REGION Network 6: IW210 - BWT Level (LT-422) - Tank #1
   RUNG wire#powerrail
      { S7_Templates := "[SrcType := Int, DestType := Real]" } Normalize(min := "20_TANKS_IP_DATA".RIO_03.FIRST_TANK.BWT_LEVEL_CNFG.RAW_MIN, value := "Tank 3P BWT Level", max := "20_TANKS_IP_DATA".RIO_03.FIRST_TANK.BWT_LEVEL_CNFG.RAW_MAX, out => "20_TANKS_IP_DATA".RIO_03.FIRST_TANK.BWT_LEVEL_CNFG.NORM)
      { S7_Templates := "[SrcType := Real, DestType := Real]" } Scale(min := "20_TANKS_IP_DATA".RIO_03.FIRST_TANK.BWT_LEVEL_CNFG.ENG_MIN, value := "IN_Level_WBT_3P", max := "20_TANKS_IP_DATA".RIO_03.FIRST_TANK.BWT_LEVEL_CNFG.ENG_MAX, out => "Tag_19")
      Move(in := "Data_From_WBT".Level_WBT_3P, out1 => "20_TANKS_IP_DATA".RIO_03.FIRST_TANK.BWT_LEVEL)
   END_RUNG
   // the same network as SCL:
   "20_TANKS_IP_DATA".RIO_03.FIRST_TANK.BWT_LEVEL_CNFG.NORM := NORM_X(MIN := "20_TANKS_IP_DATA".RIO_03.FIRST_TANK.BWT_LEVEL_CNFG.RAW_MIN, VALUE := "Tank 3P BWT Level", MAX := "20_TANKS_IP_DATA".RIO_03.FIRST_TANK.BWT_LEVEL_CNFG.RAW_MAX);
   "Tag_19" := SCALE_X(MIN := "20_TANKS_IP_DATA".RIO_03.FIRST_TANK.BWT_LEVEL_CNFG.ENG_MIN, VALUE := "IN_Level_WBT_3P", MAX := "20_TANKS_IP_DATA".RIO_03.FIRST_TANK.BWT_LEVEL_CNFG.ENG_MAX);
   "20_TANKS_IP_DATA".RIO_03.FIRST_TANK.BWT_LEVEL := "Data_From_WBT".Level_WBT_3P;
END_REGION

REGION Network 7: IW212 - BWT Level (LT-422) - Tank #2
   RUNG wire#powerrail
      { S7_Templates := "[SrcType := Int, DestType := Real]" } Normalize(min := "20_TANKS_IP_DATA".RIO_03.SECOND_TANK.BWT_LEVEL_CNFG.RAW_MIN, value := "Tank 3S BWT Level", max := "20_TANKS_IP_DATA".RIO_03.SECOND_TANK.BWT_LEVEL_CNFG.RAW_MAX, out => "20_TANKS_IP_DATA".RIO_03.SECOND_TANK.BWT_LEVEL_CNFG.NORM)
      { S7_Templates := "[SrcType := Real, DestType := Real]" } Scale(min := "20_TANKS_IP_DATA".RIO_03.SECOND_TANK.BWT_LEVEL_CNFG.ENG_MIN, value := "IN_Level_WBT_3S", max := "20_TANKS_IP_DATA".RIO_03.SECOND_TANK.BWT_LEVEL_CNFG.ENG_MAX, out => "Tag_21")
      Move(in := "Data_From_WBT".Level_WBT_3S, out1 => "20_TANKS_IP_DATA".RIO_03.SECOND_TANK.BWT_LEVEL)
   END_RUNG
   // the same network as SCL:
   "20_TANKS_IP_DATA".RIO_03.SECOND_TANK.BWT_LEVEL_CNFG.NORM := NORM_X(MIN := "20_TANKS_IP_DATA".RIO_03.SECOND_TANK.BWT_LEVEL_CNFG.RAW_MIN, VALUE := "Tank 3S BWT Level", MAX := "20_TANKS_IP_DATA".RIO_03.SECOND_TANK.BWT_LEVEL_CNFG.RAW_MAX);
   "Tag_21" := SCALE_X(MIN := "20_TANKS_IP_DATA".RIO_03.SECOND_TANK.BWT_LEVEL_CNFG.ENG_MIN, VALUE := "IN_Level_WBT_3S", MAX := "20_TANKS_IP_DATA".RIO_03.SECOND_TANK.BWT_LEVEL_CNFG.ENG_MAX);
   "20_TANKS_IP_DATA".RIO_03.SECOND_TANK.BWT_LEVEL := "Data_From_WBT".Level_WBT_3S;
END_REGION

REGION Network 8: IW214 - Spare Input - Tank #1
   RUNG wire#powerrail
      { S7_Templates := "[SrcType := Int, DestType := Real]" } Normalize(min := "20_TANKS_IP_DATA".RIO_03.FIRST_TANK.SPARE_AI_1_CNFG.RAW_MIN, value := "RIO3_SPR_AI_214", max := "20_TANKS_IP_DATA".RIO_03.FIRST_TANK.SPARE_AI_1_CNFG.RAW_MAX, out => "20_TANKS_IP_DATA".RIO_03.FIRST_TANK.SPARE_AI_1_CNFG.NORM)
      { S7_Templates := "[SrcType := Real, DestType := Real]" } Scale(min := "20_TANKS_IP_DATA".RIO_03.FIRST_TANK.SPARE_AI_1_CNFG.ENG_MIN, value := "20_TANKS_IP_DATA".RIO_03.FIRST_TANK.SPARE_AI_1_CNFG.NORM, max := "20_TANKS_IP_DATA".RIO_03.FIRST_TANK.SPARE_AI_1_CNFG.ENG_MAX, out => "20_TANKS_IP_DATA".RIO_03.FIRST_TANK.SPARE_AI_1)
   END_RUNG
   // the same network as SCL:
   "20_TANKS_IP_DATA".RIO_03.FIRST_TANK.SPARE_AI_1_CNFG.NORM := NORM_X(MIN := "20_TANKS_IP_DATA".RIO_03.FIRST_TANK.SPARE_AI_1_CNFG.RAW_MIN, VALUE := "RIO3_SPR_AI_214", MAX := "20_TANKS_IP_DATA".RIO_03.FIRST_TANK.SPARE_AI_1_CNFG.RAW_MAX);
   "20_TANKS_IP_DATA".RIO_03.FIRST_TANK.SPARE_AI_1 := SCALE_X(MIN := "20_TANKS_IP_DATA".RIO_03.FIRST_TANK.SPARE_AI_1_CNFG.ENG_MIN, VALUE := "20_TANKS_IP_DATA".RIO_03.FIRST_TANK.SPARE_AI_1_CNFG.NORM, MAX := "20_TANKS_IP_DATA".RIO_03.FIRST_TANK.SPARE_AI_1_CNFG.ENG_MAX);
END_REGION

REGION Network 9: IW216 - BWT Ph (426) - Tank #1
   RUNG wire#powerrail
      { S7_Templates := "[SrcType := Int, DestType := Real]" } Normalize(min := "20_TANKS_IP_DATA".RIO_03.FIRST_TANK.BWT_PH_CNFG.RAW_MIN, value := "Tank 3P BWT ph", max := "20_TANKS_IP_DATA".RIO_03.FIRST_TANK.BWT_PH_CNFG.RAW_MAX, out => "20_TANKS_IP_DATA".RIO_03.FIRST_TANK.BWT_PH_CNFG.NORM)
      { S7_Templates := "[SrcType := Real, DestType := Real]" } Scale(min := "20_TANKS_IP_DATA".RIO_03.FIRST_TANK.BWT_PH_CNFG.ENG_MIN, value := "20_TANKS_IP_DATA".RIO_03.FIRST_TANK.BWT_PH_CNFG.NORM, max := "20_TANKS_IP_DATA".RIO_03.FIRST_TANK.BWT_PH_CNFG.ENG_MAX, out => "20_TANKS_IP_DATA".RIO_03.FIRST_TANK.BWT_PH)
   END_RUNG
   // the same network as SCL:
   "20_TANKS_IP_DATA".RIO_03.FIRST_TANK.BWT_PH_CNFG.NORM := NORM_X(MIN := "20_TANKS_IP_DATA".RIO_03.FIRST_TANK.BWT_PH_CNFG.RAW_MIN, VALUE := "Tank 3P BWT ph", MAX := "20_TANKS_IP_DATA".RIO_03.FIRST_TANK.BWT_PH_CNFG.RAW_MAX);
   "20_TANKS_IP_DATA".RIO_03.FIRST_TANK.BWT_PH := SCALE_X(MIN := "20_TANKS_IP_DATA".RIO_03.FIRST_TANK.BWT_PH_CNFG.ENG_MIN, VALUE := "20_TANKS_IP_DATA".RIO_03.FIRST_TANK.BWT_PH_CNFG.NORM, MAX := "20_TANKS_IP_DATA".RIO_03.FIRST_TANK.BWT_PH_CNFG.ENG_MAX);
END_REGION

REGION Network 10: IW218 - BWT Temperature (426) - Tank #1
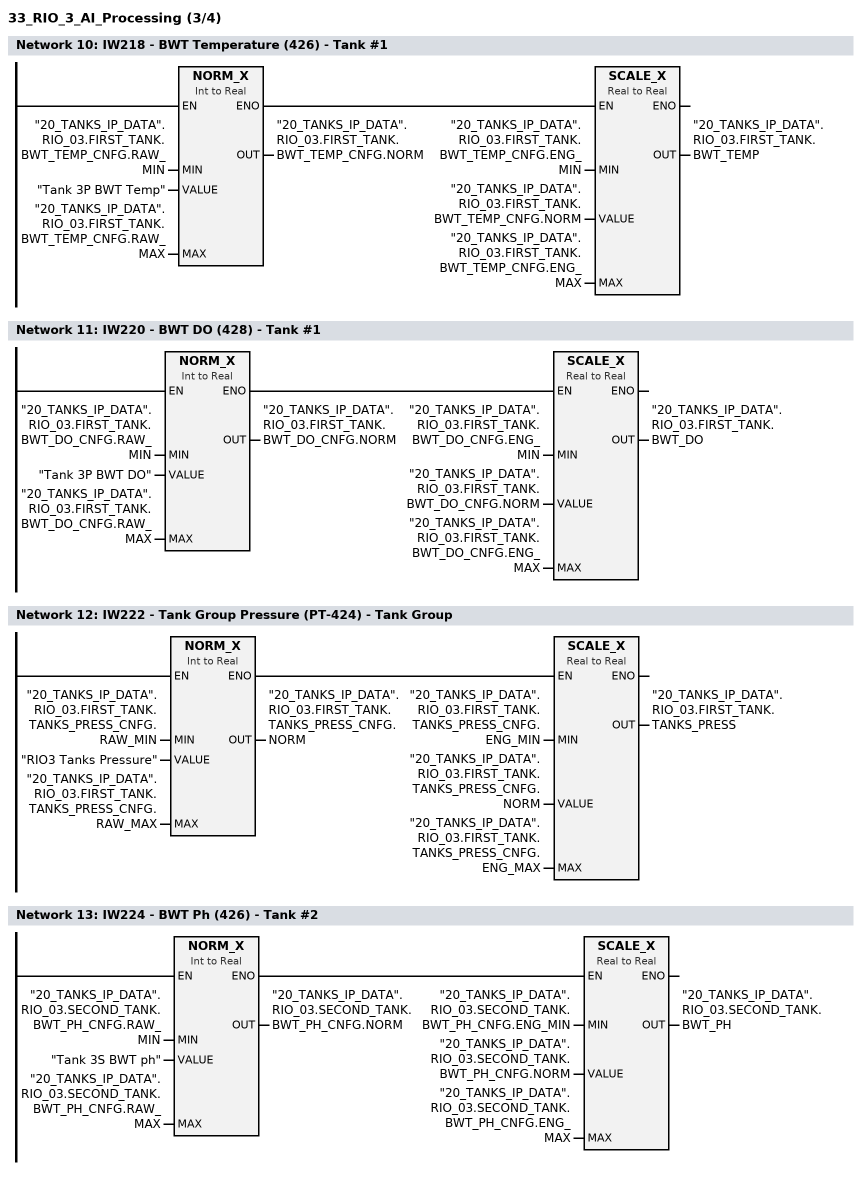
   RUNG wire#powerrail
      { S7_Templates := "[SrcType := Int, DestType := Real]" } Normalize(min := "20_TANKS_IP_DATA".RIO_03.FIRST_TANK.BWT_TEMP_CNFG.RAW_MIN, value := "Tank 3P BWT Temp", max := "20_TANKS_IP_DATA".RIO_03.FIRST_TANK.BWT_TEMP_CNFG.RAW_MAX, out => "20_TANKS_IP_DATA".RIO_03.FIRST_TANK.BWT_TEMP_CNFG.NORM)
      { S7_Templates := "[SrcType := Real, DestType := Real]" } Scale(min := "20_TANKS_IP_DATA".RIO_03.FIRST_TANK.BWT_TEMP_CNFG.ENG_MIN, value := "20_TANKS_IP_DATA".RIO_03.FIRST_TANK.BWT_TEMP_CNFG.NORM, max := "20_TANKS_IP_DATA".RIO_03.FIRST_TANK.BWT_TEMP_CNFG.ENG_MAX, out => "20_TANKS_IP_DATA".RIO_03.FIRST_TANK.BWT_TEMP)
   END_RUNG
   // the same network as SCL:
   "20_TANKS_IP_DATA".RIO_03.FIRST_TANK.BWT_TEMP_CNFG.NORM := NORM_X(MIN := "20_TANKS_IP_DATA".RIO_03.FIRST_TANK.BWT_TEMP_CNFG.RAW_MIN, VALUE := "Tank 3P BWT Temp", MAX := "20_TANKS_IP_DATA".RIO_03.FIRST_TANK.BWT_TEMP_CNFG.RAW_MAX);
   "20_TANKS_IP_DATA".RIO_03.FIRST_TANK.BWT_TEMP := SCALE_X(MIN := "20_TANKS_IP_DATA".RIO_03.FIRST_TANK.BWT_TEMP_CNFG.ENG_MIN, VALUE := "20_TANKS_IP_DATA".RIO_03.FIRST_TANK.BWT_TEMP_CNFG.NORM, MAX := "20_TANKS_IP_DATA".RIO_03.FIRST_TANK.BWT_TEMP_CNFG.ENG_MAX);
END_REGION

REGION Network 11: IW220 - BWT DO (428) - Tank #1
   RUNG wire#powerrail
      { S7_Templates := "[SrcType := Int, DestType := Real]" } Normalize(min := "20_TANKS_IP_DATA".RIO_03.FIRST_TANK.BWT_DO_CNFG.RAW_MIN, value := "Tank 3P BWT DO", max := "20_TANKS_IP_DATA".RIO_03.FIRST_TANK.BWT_DO_CNFG.RAW_MAX, out => "20_TANKS_IP_DATA".RIO_03.FIRST_TANK.BWT_DO_CNFG.NORM)
      { S7_Templates := "[SrcType := Real, DestType := Real]" } Scale(min := "20_TANKS_IP_DATA".RIO_03.FIRST_TANK.BWT_DO_CNFG.ENG_MIN, value := "20_TANKS_IP_DATA".RIO_03.FIRST_TANK.BWT_DO_CNFG.NORM, max := "20_TANKS_IP_DATA".RIO_03.FIRST_TANK.BWT_DO_CNFG.ENG_MAX, out => "20_TANKS_IP_DATA".RIO_03.FIRST_TANK.BWT_DO)
   END_RUNG
   // the same network as SCL:
   "20_TANKS_IP_DATA".RIO_03.FIRST_TANK.BWT_DO_CNFG.NORM := NORM_X(MIN := "20_TANKS_IP_DATA".RIO_03.FIRST_TANK.BWT_DO_CNFG.RAW_MIN, VALUE := "Tank 3P BWT DO", MAX := "20_TANKS_IP_DATA".RIO_03.FIRST_TANK.BWT_DO_CNFG.RAW_MAX);
   "20_TANKS_IP_DATA".RIO_03.FIRST_TANK.BWT_DO := SCALE_X(MIN := "20_TANKS_IP_DATA".RIO_03.FIRST_TANK.BWT_DO_CNFG.ENG_MIN, VALUE := "20_TANKS_IP_DATA".RIO_03.FIRST_TANK.BWT_DO_CNFG.NORM, MAX := "20_TANKS_IP_DATA".RIO_03.FIRST_TANK.BWT_DO_CNFG.ENG_MAX);
END_REGION

REGION Network 12: IW222 - Tank Group Pressure (PT-424) - Tank Group
   RUNG wire#powerrail
      { S7_Templates := "[SrcType := Int, DestType := Real]" } Normalize(min := "20_TANKS_IP_DATA".RIO_03.FIRST_TANK.TANKS_PRESS_CNFG.RAW_MIN, value := "RIO3 Tanks Pressure", max := "20_TANKS_IP_DATA".RIO_03.FIRST_TANK.TANKS_PRESS_CNFG.RAW_MAX, out => "20_TANKS_IP_DATA".RIO_03.FIRST_TANK.TANKS_PRESS_CNFG.NORM)
      { S7_Templates := "[SrcType := Real, DestType := Real]" } Scale(min := "20_TANKS_IP_DATA".RIO_03.FIRST_TANK.TANKS_PRESS_CNFG.ENG_MIN, value := "20_TANKS_IP_DATA".RIO_03.FIRST_TANK.TANKS_PRESS_CNFG.NORM, max := "20_TANKS_IP_DATA".RIO_03.FIRST_TANK.TANKS_PRESS_CNFG.ENG_MAX, out => "20_TANKS_IP_DATA".RIO_03.FIRST_TANK.TANKS_PRESS)
   END_RUNG
   // the same network as SCL:
   "20_TANKS_IP_DATA".RIO_03.FIRST_TANK.TANKS_PRESS_CNFG.NORM := NORM_X(MIN := "20_TANKS_IP_DATA".RIO_03.FIRST_TANK.TANKS_PRESS_CNFG.RAW_MIN, VALUE := "RIO3 Tanks Pressure", MAX := "20_TANKS_IP_DATA".RIO_03.FIRST_TANK.TANKS_PRESS_CNFG.RAW_MAX);
   "20_TANKS_IP_DATA".RIO_03.FIRST_TANK.TANKS_PRESS := SCALE_X(MIN := "20_TANKS_IP_DATA".RIO_03.FIRST_TANK.TANKS_PRESS_CNFG.ENG_MIN, VALUE := "20_TANKS_IP_DATA".RIO_03.FIRST_TANK.TANKS_PRESS_CNFG.NORM, MAX := "20_TANKS_IP_DATA".RIO_03.FIRST_TANK.TANKS_PRESS_CNFG.ENG_MAX);
END_REGION

REGION Network 13: IW224 - BWT Ph (426) - Tank #2
   RUNG wire#powerrail
      { S7_Templates := "[SrcType := Int, DestType := Real]" } Normalize(min := "20_TANKS_IP_DATA".RIO_03.SECOND_TANK.BWT_PH_CNFG.RAW_MIN, value := "Tank 3S BWT ph", max := "20_TANKS_IP_DATA".RIO_03.SECOND_TANK.BWT_PH_CNFG.RAW_MAX, out => "20_TANKS_IP_DATA".RIO_03.SECOND_TANK.BWT_PH_CNFG.NORM)
      { S7_Templates := "[SrcType := Real, DestType := Real]" } Scale(min := "20_TANKS_IP_DATA".RIO_03.SECOND_TANK.BWT_PH_CNFG.ENG_MIN, value := "20_TANKS_IP_DATA".RIO_03.SECOND_TANK.BWT_PH_CNFG.NORM, max := "20_TANKS_IP_DATA".RIO_03.SECOND_TANK.BWT_PH_CNFG.ENG_MAX, out => "20_TANKS_IP_DATA".RIO_03.SECOND_TANK.BWT_PH)
   END_RUNG
   // the same network as SCL:
   "20_TANKS_IP_DATA".RIO_03.SECOND_TANK.BWT_PH_CNFG.NORM := NORM_X(MIN := "20_TANKS_IP_DATA".RIO_03.SECOND_TANK.BWT_PH_CNFG.RAW_MIN, VALUE := "Tank 3S BWT ph", MAX := "20_TANKS_IP_DATA".RIO_03.SECOND_TANK.BWT_PH_CNFG.RAW_MAX);
   "20_TANKS_IP_DATA".RIO_03.SECOND_TANK.BWT_PH := SCALE_X(MIN := "20_TANKS_IP_DATA".RIO_03.SECOND_TANK.BWT_PH_CNFG.ENG_MIN, VALUE := "20_TANKS_IP_DATA".RIO_03.SECOND_TANK.BWT_PH_CNFG.NORM, MAX := "20_TANKS_IP_DATA".RIO_03.SECOND_TANK.BWT_PH_CNFG.ENG_MAX);
END_REGION

REGION Network 14: IW226 - BWT Temperature (426) - Tank #2
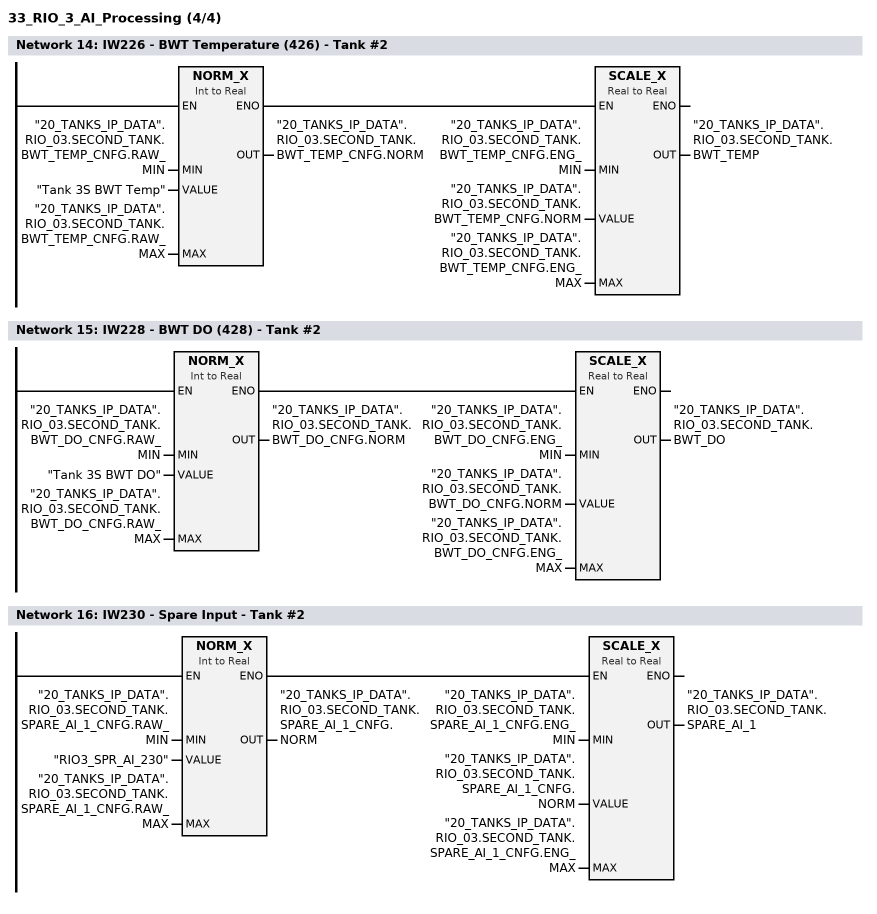
   RUNG wire#powerrail
      { S7_Templates := "[SrcType := Int, DestType := Real]" } Normalize(min := "20_TANKS_IP_DATA".RIO_03.SECOND_TANK.BWT_TEMP_CNFG.RAW_MIN, value := "Tank 3S BWT Temp", max := "20_TANKS_IP_DATA".RIO_03.SECOND_TANK.BWT_TEMP_CNFG.RAW_MAX, out => "20_TANKS_IP_DATA".RIO_03.SECOND_TANK.BWT_TEMP_CNFG.NORM)
      { S7_Templates := "[SrcType := Real, DestType := Real]" } Scale(min := "20_TANKS_IP_DATA".RIO_03.SECOND_TANK.BWT_TEMP_CNFG.ENG_MIN, value := "20_TANKS_IP_DATA".RIO_03.SECOND_TANK.BWT_TEMP_CNFG.NORM, max := "20_TANKS_IP_DATA".RIO_03.SECOND_TANK.BWT_TEMP_CNFG.ENG_MAX, out => "20_TANKS_IP_DATA".RIO_03.SECOND_TANK.BWT_TEMP)
   END_RUNG
   // the same network as SCL:
   "20_TANKS_IP_DATA".RIO_03.SECOND_TANK.BWT_TEMP_CNFG.NORM := NORM_X(MIN := "20_TANKS_IP_DATA".RIO_03.SECOND_TANK.BWT_TEMP_CNFG.RAW_MIN, VALUE := "Tank 3S BWT Temp", MAX := "20_TANKS_IP_DATA".RIO_03.SECOND_TANK.BWT_TEMP_CNFG.RAW_MAX);
   "20_TANKS_IP_DATA".RIO_03.SECOND_TANK.BWT_TEMP := SCALE_X(MIN := "20_TANKS_IP_DATA".RIO_03.SECOND_TANK.BWT_TEMP_CNFG.ENG_MIN, VALUE := "20_TANKS_IP_DATA".RIO_03.SECOND_TANK.BWT_TEMP_CNFG.NORM, MAX := "20_TANKS_IP_DATA".RIO_03.SECOND_TANK.BWT_TEMP_CNFG.ENG_MAX);
END_REGION

REGION Network 15: IW228 - BWT DO (428) - Tank #2
   RUNG wire#powerrail
      { S7_Templates := "[SrcType := Int, DestType := Real]" } Normalize(min := "20_TANKS_IP_DATA".RIO_03.SECOND_TANK.BWT_DO_CNFG.RAW_MIN, value := "Tank 3S BWT DO", max := "20_TANKS_IP_DATA".RIO_03.SECOND_TANK.BWT_DO_CNFG.RAW_MAX, out => "20_TANKS_IP_DATA".RIO_03.SECOND_TANK.BWT_DO_CNFG.NORM)
      { S7_Templates := "[SrcType := Real, DestType := Real]" } Scale(min := "20_TANKS_IP_DATA".RIO_03.SECOND_TANK.BWT_DO_CNFG.ENG_MIN, value := "20_TANKS_IP_DATA".RIO_03.SECOND_TANK.BWT_DO_CNFG.NORM, max := "20_TANKS_IP_DATA".RIO_03.SECOND_TANK.BWT_DO_CNFG.ENG_MAX, out => "20_TANKS_IP_DATA".RIO_03.SECOND_TANK.BWT_DO)
   END_RUNG
   // the same network as SCL:
   "20_TANKS_IP_DATA".RIO_03.SECOND_TANK.BWT_DO_CNFG.NORM := NORM_X(MIN := "20_TANKS_IP_DATA".RIO_03.SECOND_TANK.BWT_DO_CNFG.RAW_MIN, VALUE := "Tank 3S BWT DO", MAX := "20_TANKS_IP_DATA".RIO_03.SECOND_TANK.BWT_DO_CNFG.RAW_MAX);
   "20_TANKS_IP_DATA".RIO_03.SECOND_TANK.BWT_DO := SCALE_X(MIN := "20_TANKS_IP_DATA".RIO_03.SECOND_TANK.BWT_DO_CNFG.ENG_MIN, VALUE := "20_TANKS_IP_DATA".RIO_03.SECOND_TANK.BWT_DO_CNFG.NORM, MAX := "20_TANKS_IP_DATA".RIO_03.SECOND_TANK.BWT_DO_CNFG.ENG_MAX);
END_REGION

REGION Network 16: IW230 - Spare Input - Tank #2
   RUNG wire#powerrail
      { S7_Templates := "[SrcType := Int, DestType := Real]" } Normalize(min := "20_TANKS_IP_DATA".RIO_03.SECOND_TANK.SPARE_AI_1_CNFG.RAW_MIN, value := "RIO3_SPR_AI_230", max := "20_TANKS_IP_DATA".RIO_03.SECOND_TANK.SPARE_AI_1_CNFG.RAW_MAX, out => "20_TANKS_IP_DATA".RIO_03.SECOND_TANK.SPARE_AI_1_CNFG.NORM)
      { S7_Templates := "[SrcType := Real, DestType := Real]" } Scale(min := "20_TANKS_IP_DATA".RIO_03.SECOND_TANK.SPARE_AI_1_CNFG.ENG_MIN, value := "20_TANKS_IP_DATA".RIO_03.SECOND_TANK.SPARE_AI_1_CNFG.NORM, max := "20_TANKS_IP_DATA".RIO_03.SECOND_TANK.SPARE_AI_1_CNFG.ENG_MAX, out => "20_TANKS_IP_DATA".RIO_03.SECOND_TANK.SPARE_AI_1)
   END_RUNG
   // the same network as SCL:
   "20_TANKS_IP_DATA".RIO_03.SECOND_TANK.SPARE_AI_1_CNFG.NORM := NORM_X(MIN := "20_TANKS_IP_DATA".RIO_03.SECOND_TANK.SPARE_AI_1_CNFG.RAW_MIN, VALUE := "RIO3_SPR_AI_230", MAX := "20_TANKS_IP_DATA".RIO_03.SECOND_TANK.SPARE_AI_1_CNFG.RAW_MAX);
   "20_TANKS_IP_DATA".RIO_03.SECOND_TANK.SPARE_AI_1 := SCALE_X(MIN := "20_TANKS_IP_DATA".RIO_03.SECOND_TANK.SPARE_AI_1_CNFG.ENG_MIN, VALUE := "20_TANKS_IP_DATA".RIO_03.SECOND_TANK.SPARE_AI_1_CNFG.NORM, MAX := "20_TANKS_IP_DATA".RIO_03.SECOND_TANK.SPARE_AI_1_CNFG.ENG_MAX);
END_REGION
END_FUNCTION

FUNCTION "34_RIO_4_AI_Processing" : Void   // FC34, LAD
TITLE = Analogue Input Processing (Tank 1 = 4P, Tank 2 = 4S)
{ S7_Optimized_Access := 'TRUE' }
AUTHOR : JRS
VERSION : 0.1
// To process raw inputs prior to code use
BEGIN

REGION Network 1: IW260 - USD Flow (FIT-418) - Tank #1
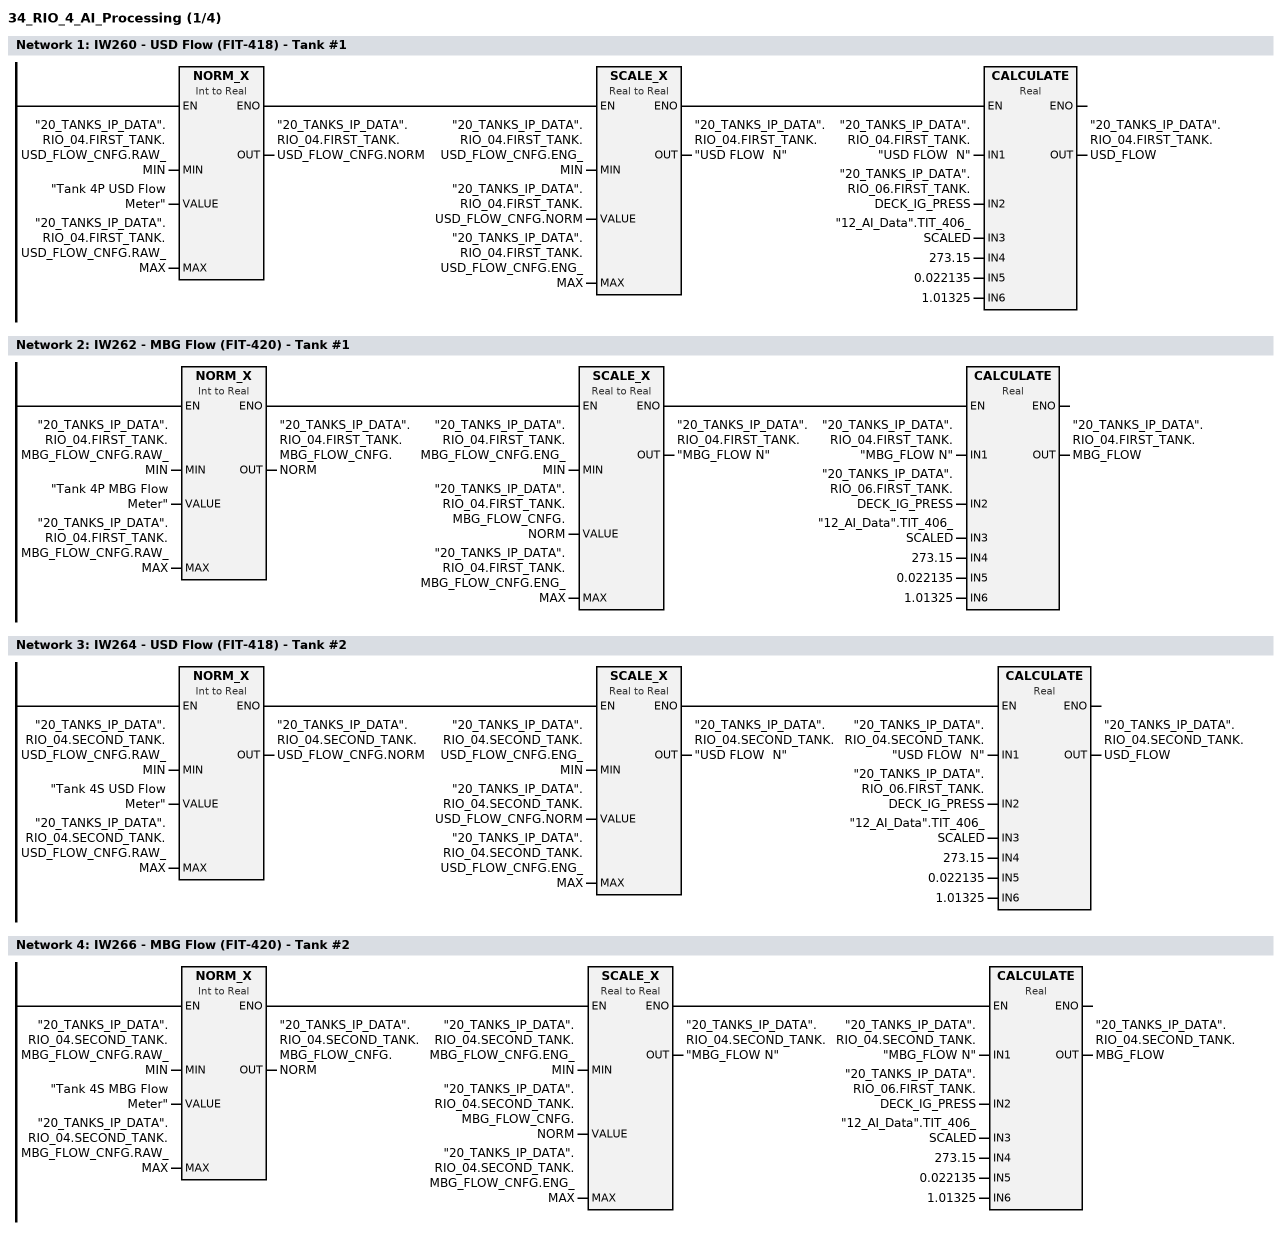
   RUNG wire#powerrail
      { S7_Templates := "[SrcType := Int, DestType := Real]" } Normalize(min := "20_TANKS_IP_DATA".RIO_04.FIRST_TANK.USD_FLOW_CNFG.RAW_MIN, value := "Tank 4P USD Flow Meter", max := "20_TANKS_IP_DATA".RIO_04.FIRST_TANK.USD_FLOW_CNFG.RAW_MAX, out => "20_TANKS_IP_DATA".RIO_04.FIRST_TANK.USD_FLOW_CNFG.NORM)
      { S7_Templates := "[SrcType := Real, DestType := Real]" } Scale(min := "20_TANKS_IP_DATA".RIO_04.FIRST_TANK.USD_FLOW_CNFG.ENG_MIN, value := "20_TANKS_IP_DATA".RIO_04.FIRST_TANK.USD_FLOW_CNFG.NORM, max := "20_TANKS_IP_DATA".RIO_04.FIRST_TANK.USD_FLOW_CNFG.ENG_MAX, out => "20_TANKS_IP_DATA".RIO_04.FIRST_TANK."USD FLOW  N")
      { S7_Templates := "SrcType := Real"; S7_Expression := "IN1*(IN2+IN6)/IN6*IN4/(IN3+IN4)" } Calculate(in1 := "20_TANKS_IP_DATA".RIO_04.FIRST_TANK."USD FLOW  N", in2 := "20_TANKS_IP_DATA".RIO_06.FIRST_TANK.DECK_IG_PRESS, in3 := "12_AI_Data".TIT_406_SCALED, in4 := 273.15, in5 := 0.022135, in6 := 1.01325, out => "20_TANKS_IP_DATA".RIO_04.FIRST_TANK.USD_FLOW)
   END_RUNG
   // the same network as SCL:
   "20_TANKS_IP_DATA".RIO_04.FIRST_TANK.USD_FLOW_CNFG.NORM := NORM_X(MIN := "20_TANKS_IP_DATA".RIO_04.FIRST_TANK.USD_FLOW_CNFG.RAW_MIN, VALUE := "Tank 4P USD Flow Meter", MAX := "20_TANKS_IP_DATA".RIO_04.FIRST_TANK.USD_FLOW_CNFG.RAW_MAX);
   "20_TANKS_IP_DATA".RIO_04.FIRST_TANK."USD FLOW  N" := SCALE_X(MIN := "20_TANKS_IP_DATA".RIO_04.FIRST_TANK.USD_FLOW_CNFG.ENG_MIN, VALUE := "20_TANKS_IP_DATA".RIO_04.FIRST_TANK.USD_FLOW_CNFG.NORM, MAX := "20_TANKS_IP_DATA".RIO_04.FIRST_TANK.USD_FLOW_CNFG.ENG_MAX);
   "20_TANKS_IP_DATA".RIO_04.FIRST_TANK.USD_FLOW := "20_TANKS_IP_DATA".RIO_04.FIRST_TANK."USD FLOW  N"*("20_TANKS_IP_DATA".RIO_06.FIRST_TANK.DECK_IG_PRESS+1.01325)/1.01325*273.15/("12_AI_Data".TIT_406_SCALED+273.15);
END_REGION

REGION Network 2: IW262 - MBG Flow (FIT-420) - Tank #1
   RUNG wire#powerrail
      { S7_Templates := "[SrcType := Int, DestType := Real]" } Normalize(min := "20_TANKS_IP_DATA".RIO_04.FIRST_TANK.MBG_FLOW_CNFG.RAW_MIN, value := "Tank 4P MBG Flow Meter", max := "20_TANKS_IP_DATA".RIO_04.FIRST_TANK.MBG_FLOW_CNFG.RAW_MAX, out => "20_TANKS_IP_DATA".RIO_04.FIRST_TANK.MBG_FLOW_CNFG.NORM)
      { S7_Templates := "[SrcType := Real, DestType := Real]" } Scale(min := "20_TANKS_IP_DATA".RIO_04.FIRST_TANK.MBG_FLOW_CNFG.ENG_MIN, value := "20_TANKS_IP_DATA".RIO_04.FIRST_TANK.MBG_FLOW_CNFG.NORM, max := "20_TANKS_IP_DATA".RIO_04.FIRST_TANK.MBG_FLOW_CNFG.ENG_MAX, out => "20_TANKS_IP_DATA".RIO_04.FIRST_TANK."MBG_FLOW N")
      { S7_Templates := "SrcType := Real"; S7_Expression := "IN1*(IN2+IN6)/IN6*IN4/(IN3+IN4)" } Calculate(in1 := "20_TANKS_IP_DATA".RIO_04.FIRST_TANK."MBG_FLOW N", in2 := "20_TANKS_IP_DATA".RIO_06.FIRST_TANK.DECK_IG_PRESS, in3 := "12_AI_Data".TIT_406_SCALED, in4 := 273.15, in5 := 0.022135, in6 := 1.01325, out => "20_TANKS_IP_DATA".RIO_04.FIRST_TANK.MBG_FLOW)
   END_RUNG
   // the same network as SCL:
   "20_TANKS_IP_DATA".RIO_04.FIRST_TANK.MBG_FLOW_CNFG.NORM := NORM_X(MIN := "20_TANKS_IP_DATA".RIO_04.FIRST_TANK.MBG_FLOW_CNFG.RAW_MIN, VALUE := "Tank 4P MBG Flow Meter", MAX := "20_TANKS_IP_DATA".RIO_04.FIRST_TANK.MBG_FLOW_CNFG.RAW_MAX);
   "20_TANKS_IP_DATA".RIO_04.FIRST_TANK."MBG_FLOW N" := SCALE_X(MIN := "20_TANKS_IP_DATA".RIO_04.FIRST_TANK.MBG_FLOW_CNFG.ENG_MIN, VALUE := "20_TANKS_IP_DATA".RIO_04.FIRST_TANK.MBG_FLOW_CNFG.NORM, MAX := "20_TANKS_IP_DATA".RIO_04.FIRST_TANK.MBG_FLOW_CNFG.ENG_MAX);
   "20_TANKS_IP_DATA".RIO_04.FIRST_TANK.MBG_FLOW := "20_TANKS_IP_DATA".RIO_04.FIRST_TANK."MBG_FLOW N"*("20_TANKS_IP_DATA".RIO_06.FIRST_TANK.DECK_IG_PRESS+1.01325)/1.01325*273.15/("12_AI_Data".TIT_406_SCALED+273.15);
END_REGION

REGION Network 3: IW264 - USD Flow (FIT-418) - Tank #2
   RUNG wire#powerrail
      { S7_Templates := "[SrcType := Int, DestType := Real]" } Normalize(min := "20_TANKS_IP_DATA".RIO_04.SECOND_TANK.USD_FLOW_CNFG.RAW_MIN, value := "Tank 4S USD Flow Meter", max := "20_TANKS_IP_DATA".RIO_04.SECOND_TANK.USD_FLOW_CNFG.RAW_MAX, out => "20_TANKS_IP_DATA".RIO_04.SECOND_TANK.USD_FLOW_CNFG.NORM)
      { S7_Templates := "[SrcType := Real, DestType := Real]" } Scale(min := "20_TANKS_IP_DATA".RIO_04.SECOND_TANK.USD_FLOW_CNFG.ENG_MIN, value := "20_TANKS_IP_DATA".RIO_04.SECOND_TANK.USD_FLOW_CNFG.NORM, max := "20_TANKS_IP_DATA".RIO_04.SECOND_TANK.USD_FLOW_CNFG.ENG_MAX, out => "20_TANKS_IP_DATA".RIO_04.SECOND_TANK."USD FLOW  N")
      { S7_Templates := "SrcType := Real"; S7_Expression := "IN1*(IN2+IN6)/IN6*IN4/(IN3+IN4)" } Calculate(in1 := "20_TANKS_IP_DATA".RIO_04.SECOND_TANK."USD FLOW  N", in2 := "20_TANKS_IP_DATA".RIO_06.FIRST_TANK.DECK_IG_PRESS, in3 := "12_AI_Data".TIT_406_SCALED, in4 := 273.15, in5 := 0.022135, in6 := 1.01325, out => "20_TANKS_IP_DATA".RIO_04.SECOND_TANK.USD_FLOW)
   END_RUNG
   // the same network as SCL:
   "20_TANKS_IP_DATA".RIO_04.SECOND_TANK.USD_FLOW_CNFG.NORM := NORM_X(MIN := "20_TANKS_IP_DATA".RIO_04.SECOND_TANK.USD_FLOW_CNFG.RAW_MIN, VALUE := "Tank 4S USD Flow Meter", MAX := "20_TANKS_IP_DATA".RIO_04.SECOND_TANK.USD_FLOW_CNFG.RAW_MAX);
   "20_TANKS_IP_DATA".RIO_04.SECOND_TANK."USD FLOW  N" := SCALE_X(MIN := "20_TANKS_IP_DATA".RIO_04.SECOND_TANK.USD_FLOW_CNFG.ENG_MIN, VALUE := "20_TANKS_IP_DATA".RIO_04.SECOND_TANK.USD_FLOW_CNFG.NORM, MAX := "20_TANKS_IP_DATA".RIO_04.SECOND_TANK.USD_FLOW_CNFG.ENG_MAX);
   "20_TANKS_IP_DATA".RIO_04.SECOND_TANK.USD_FLOW := "20_TANKS_IP_DATA".RIO_04.SECOND_TANK."USD FLOW  N"*("20_TANKS_IP_DATA".RIO_06.FIRST_TANK.DECK_IG_PRESS+1.01325)/1.01325*273.15/("12_AI_Data".TIT_406_SCALED+273.15);
END_REGION

REGION Network 4: IW266 - MBG Flow (FIT-420) - Tank #2
   RUNG wire#powerrail
      { S7_Templates := "[SrcType := Int, DestType := Real]" } Normalize(min := "20_TANKS_IP_DATA".RIO_04.SECOND_TANK.MBG_FLOW_CNFG.RAW_MIN, value := "Tank 4S MBG Flow Meter", max := "20_TANKS_IP_DATA".RIO_04.SECOND_TANK.MBG_FLOW_CNFG.RAW_MAX, out => "20_TANKS_IP_DATA".RIO_04.SECOND_TANK.MBG_FLOW_CNFG.NORM)
      { S7_Templates := "[SrcType := Real, DestType := Real]" } Scale(min := "20_TANKS_IP_DATA".RIO_04.SECOND_TANK.MBG_FLOW_CNFG.ENG_MIN, value := "20_TANKS_IP_DATA".RIO_04.SECOND_TANK.MBG_FLOW_CNFG.NORM, max := "20_TANKS_IP_DATA".RIO_04.SECOND_TANK.MBG_FLOW_CNFG.ENG_MAX, out => "20_TANKS_IP_DATA".RIO_04.SECOND_TANK."MBG_FLOW N")
      { S7_Templates := "SrcType := Real"; S7_Expression := "IN1*(IN2+IN6)/IN6*IN4/(IN3+IN4)" } Calculate(in1 := "20_TANKS_IP_DATA".RIO_04.SECOND_TANK."MBG_FLOW N", in2 := "20_TANKS_IP_DATA".RIO_06.FIRST_TANK.DECK_IG_PRESS, in3 := "12_AI_Data".TIT_406_SCALED, in4 := 273.15, in5 := 0.022135, in6 := 1.01325, out => "20_TANKS_IP_DATA".RIO_04.SECOND_TANK.MBG_FLOW)
   END_RUNG
   // the same network as SCL:
   "20_TANKS_IP_DATA".RIO_04.SECOND_TANK.MBG_FLOW_CNFG.NORM := NORM_X(MIN := "20_TANKS_IP_DATA".RIO_04.SECOND_TANK.MBG_FLOW_CNFG.RAW_MIN, VALUE := "Tank 4S MBG Flow Meter", MAX := "20_TANKS_IP_DATA".RIO_04.SECOND_TANK.MBG_FLOW_CNFG.RAW_MAX);
   "20_TANKS_IP_DATA".RIO_04.SECOND_TANK."MBG_FLOW N" := SCALE_X(MIN := "20_TANKS_IP_DATA".RIO_04.SECOND_TANK.MBG_FLOW_CNFG.ENG_MIN, VALUE := "20_TANKS_IP_DATA".RIO_04.SECOND_TANK.MBG_FLOW_CNFG.NORM, MAX := "20_TANKS_IP_DATA".RIO_04.SECOND_TANK.MBG_FLOW_CNFG.ENG_MAX);
   "20_TANKS_IP_DATA".RIO_04.SECOND_TANK.MBG_FLOW := "20_TANKS_IP_DATA".RIO_04.SECOND_TANK."MBG_FLOW N"*("20_TANKS_IP_DATA".RIO_06.FIRST_TANK.DECK_IG_PRESS+1.01325)/1.01325*273.15/("12_AI_Data".TIT_406_SCALED+273.15);
END_REGION

REGION Network 5: IW268 - Deck Main IG Pressure (PT-415) - Tank Group
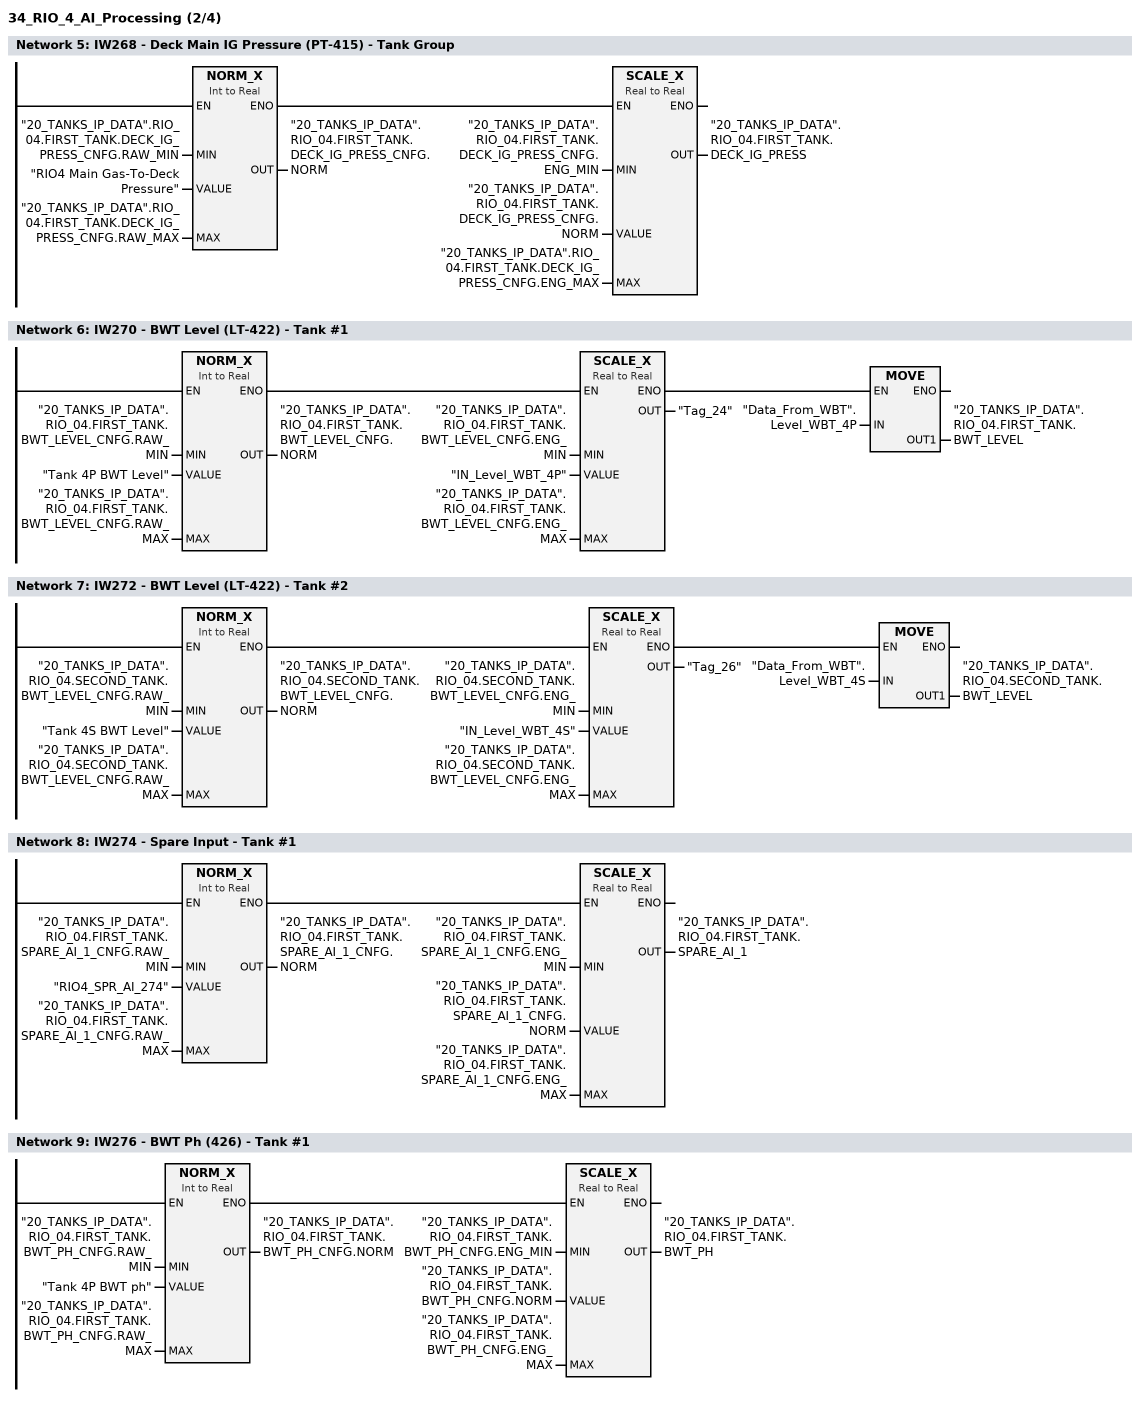
   RUNG wire#powerrail
      { S7_Templates := "[SrcType := Int, DestType := Real]" } Normalize(min := "20_TANKS_IP_DATA".RIO_04.FIRST_TANK.DECK_IG_PRESS_CNFG.RAW_MIN, value := "RIO4 Main Gas-To-Deck Pressure", max := "20_TANKS_IP_DATA".RIO_04.FIRST_TANK.DECK_IG_PRESS_CNFG.RAW_MAX, out => "20_TANKS_IP_DATA".RIO_04.FIRST_TANK.DECK_IG_PRESS_CNFG.NORM)
      { S7_Templates := "[SrcType := Real, DestType := Real]" } Scale(min := "20_TANKS_IP_DATA".RIO_04.FIRST_TANK.DECK_IG_PRESS_CNFG.ENG_MIN, value := "20_TANKS_IP_DATA".RIO_04.FIRST_TANK.DECK_IG_PRESS_CNFG.NORM, max := "20_TANKS_IP_DATA".RIO_04.FIRST_TANK.DECK_IG_PRESS_CNFG.ENG_MAX, out => "20_TANKS_IP_DATA".RIO_04.FIRST_TANK.DECK_IG_PRESS)
   END_RUNG
   // the same network as SCL:
   "20_TANKS_IP_DATA".RIO_04.FIRST_TANK.DECK_IG_PRESS_CNFG.NORM := NORM_X(MIN := "20_TANKS_IP_DATA".RIO_04.FIRST_TANK.DECK_IG_PRESS_CNFG.RAW_MIN, VALUE := "RIO4 Main Gas-To-Deck Pressure", MAX := "20_TANKS_IP_DATA".RIO_04.FIRST_TANK.DECK_IG_PRESS_CNFG.RAW_MAX);
   "20_TANKS_IP_DATA".RIO_04.FIRST_TANK.DECK_IG_PRESS := SCALE_X(MIN := "20_TANKS_IP_DATA".RIO_04.FIRST_TANK.DECK_IG_PRESS_CNFG.ENG_MIN, VALUE := "20_TANKS_IP_DATA".RIO_04.FIRST_TANK.DECK_IG_PRESS_CNFG.NORM, MAX := "20_TANKS_IP_DATA".RIO_04.FIRST_TANK.DECK_IG_PRESS_CNFG.ENG_MAX);
END_REGION

REGION Network 6: IW270 - BWT Level (LT-422) - Tank #1
   RUNG wire#powerrail
      { S7_Templates := "[SrcType := Int, DestType := Real]" } Normalize(min := "20_TANKS_IP_DATA".RIO_04.FIRST_TANK.BWT_LEVEL_CNFG.RAW_MIN, value := "Tank 4P BWT Level", max := "20_TANKS_IP_DATA".RIO_04.FIRST_TANK.BWT_LEVEL_CNFG.RAW_MAX, out => "20_TANKS_IP_DATA".RIO_04.FIRST_TANK.BWT_LEVEL_CNFG.NORM)
      { S7_Templates := "[SrcType := Real, DestType := Real]" } Scale(min := "20_TANKS_IP_DATA".RIO_04.FIRST_TANK.BWT_LEVEL_CNFG.ENG_MIN, value := "IN_Level_WBT_4P", max := "20_TANKS_IP_DATA".RIO_04.FIRST_TANK.BWT_LEVEL_CNFG.ENG_MAX, out => "Tag_24")
      Move(in := "Data_From_WBT".Level_WBT_4P, out1 => "20_TANKS_IP_DATA".RIO_04.FIRST_TANK.BWT_LEVEL)
   END_RUNG
   // the same network as SCL:
   "20_TANKS_IP_DATA".RIO_04.FIRST_TANK.BWT_LEVEL_CNFG.NORM := NORM_X(MIN := "20_TANKS_IP_DATA".RIO_04.FIRST_TANK.BWT_LEVEL_CNFG.RAW_MIN, VALUE := "Tank 4P BWT Level", MAX := "20_TANKS_IP_DATA".RIO_04.FIRST_TANK.BWT_LEVEL_CNFG.RAW_MAX);
   "Tag_24" := SCALE_X(MIN := "20_TANKS_IP_DATA".RIO_04.FIRST_TANK.BWT_LEVEL_CNFG.ENG_MIN, VALUE := "IN_Level_WBT_4P", MAX := "20_TANKS_IP_DATA".RIO_04.FIRST_TANK.BWT_LEVEL_CNFG.ENG_MAX);
   "20_TANKS_IP_DATA".RIO_04.FIRST_TANK.BWT_LEVEL := "Data_From_WBT".Level_WBT_4P;
END_REGION
